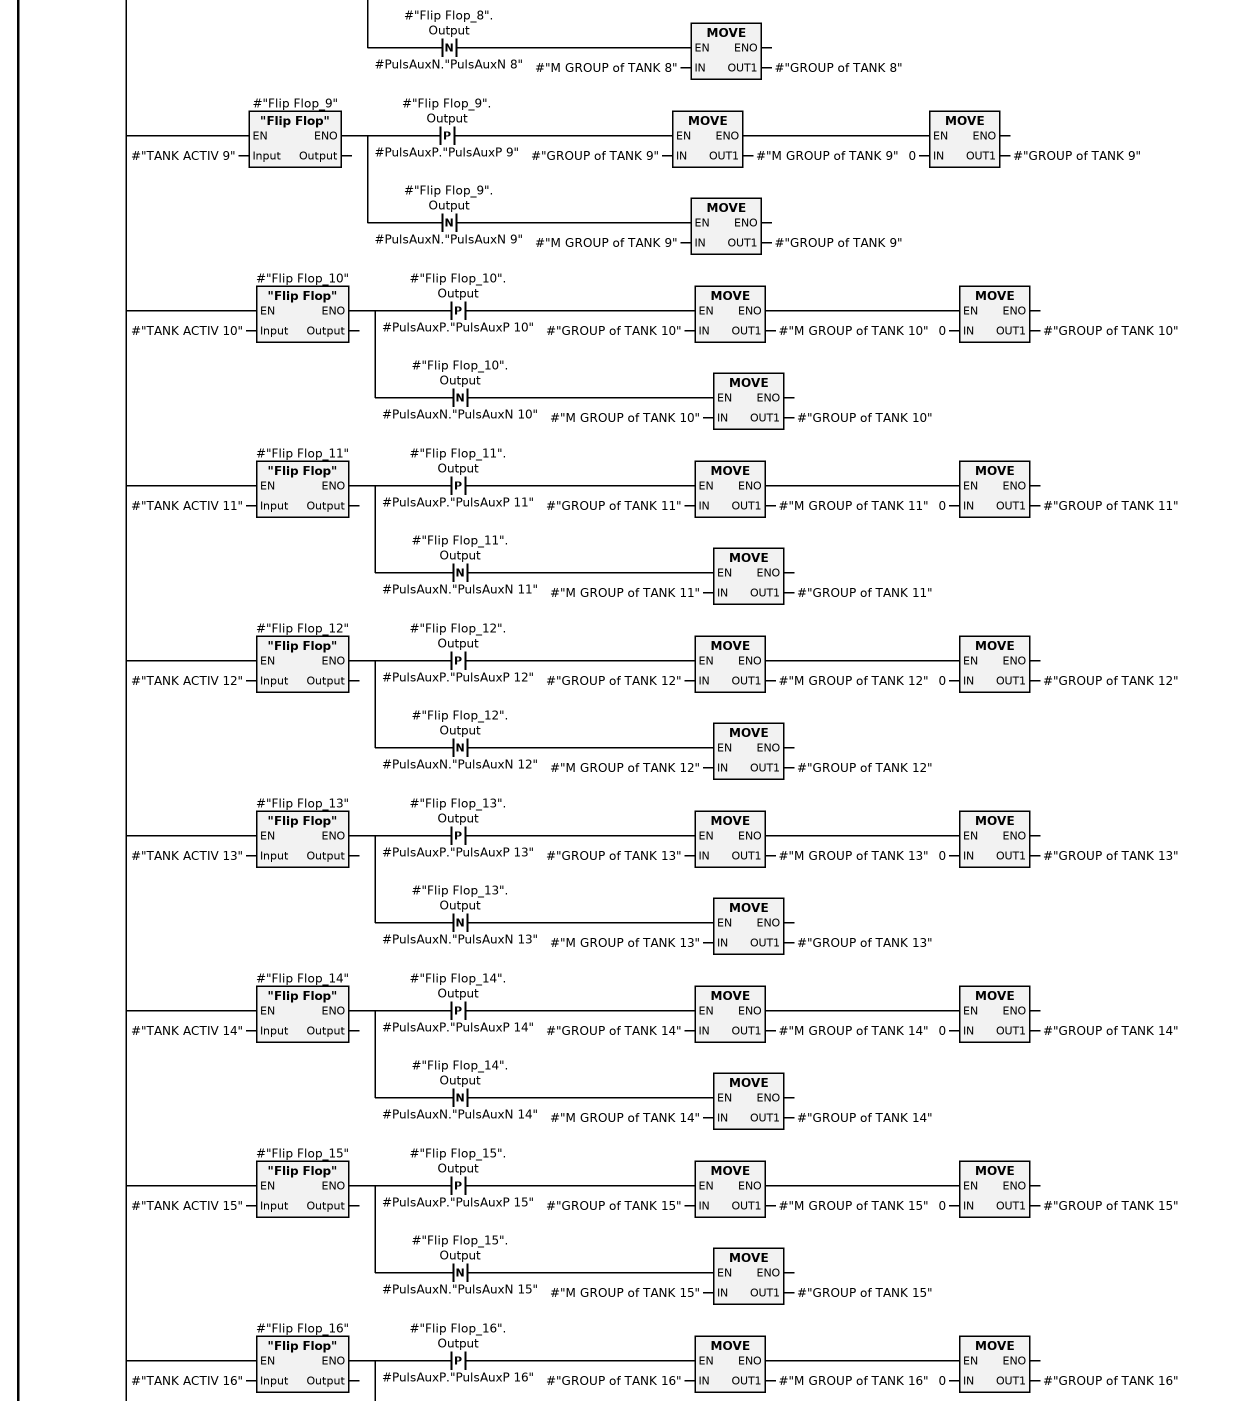
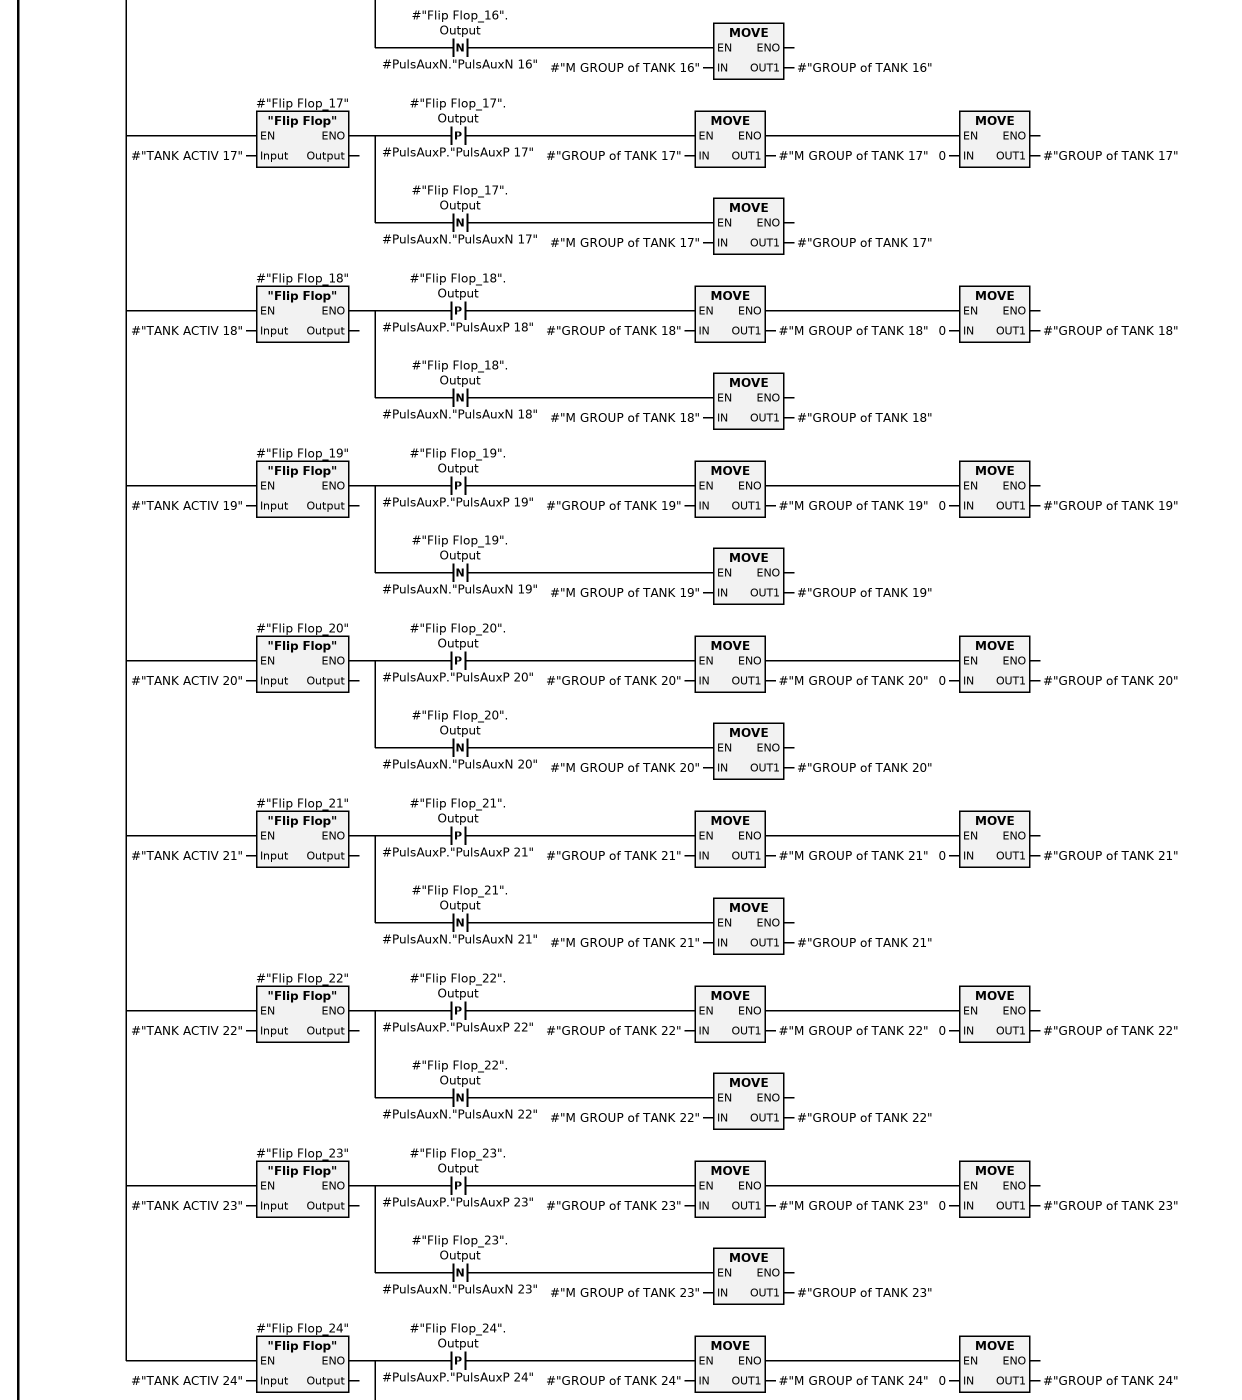
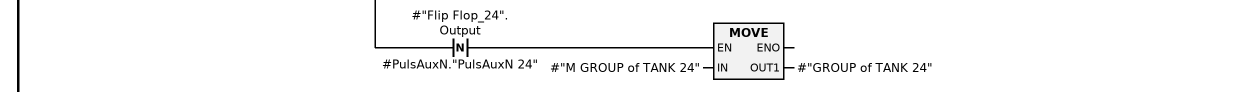
   RUNG wire#powerrail
      I_Contact( #SetGroupSR )
      wire#w1
      #"Flip Flop_1"(Input := #"TANK ACTIV 1", Output =>)
      wire#w2
      P_Contact(operand := #"Flip Flop_1".Output, bit := #PulsAuxP."PulsAuxP 1")
      Move(in := #"GROUP of TANK 1", out1 => #"M GROUP of TANK 1")
      Move(in := 0, out1 => #"GROUP of TANK 1")
   END_RUNG
   RUNG wire#w2
      N_Contact(operand := #"Flip Flop_1".Output, bit := #PulsAuxN."PulsAuxN 1")
      Move(in := #"M GROUP of TANK 1", out1 => #"GROUP of TANK 1")
   END_RUNG
   RUNG wire#w1
      #"Flip Flop_2"(Input := #"TANK ACTIV 2", Output =>)
      wire#w3
      P_Contact(operand := #"Flip Flop_2".Output, bit := #PulsAuxP."PulsAuxP 2")
      Move(in := #"GROUP of TANK 2", out1 => #"M GROUP of TANK 2")
      Move(in := 0, out1 => #"GROUP of TANK 2")
   END_RUNG
   RUNG wire#w3
      N_Contact(operand := #"Flip Flop_2".Output, bit := #PulsAuxN."PulsAuxN 2")
      Move(in := #"M GROUP of TANK 2", out1 => #"GROUP of TANK 2")
   END_RUNG
   RUNG wire#w1
      #"Flip Flop_3"(Input := #"TANK ACTIV 3", Output =>)
      wire#w4
      P_Contact(operand := #"Flip Flop_3".Output, bit := #PulsAuxP."PulsAuxP 3")
      Move(in := #"GROUP of TANK 3", out1 => #"M GROUP of TANK 3")
      Move(in := 0, out1 => #"GROUP of TANK 3")
   END_RUNG
   RUNG wire#w4
      N_Contact(operand := #"Flip Flop_3".Output, bit := #PulsAuxN."PulsAuxN 3")
      Move(in := #"M GROUP of TANK 3", out1 => #"GROUP of TANK 3")
   END_RUNG
   RUNG wire#w1
      #"Flip Flop_4"(Input := #"TANK ACTIV 4", Output =>)
      wire#w5
      P_Contact(operand := #"Flip Flop_4".Output, bit := #PulsAuxP."PulsAuxP 4")
      Move(in := #"GROUP of TANK 4", out1 => #"M GROUP of TANK 4")
      Move(in := 0, out1 => #"GROUP of TANK 4")
   END_RUNG
   RUNG wire#w5
      N_Contact(operand := #"Flip Flop_4".Output, bit := #PulsAuxN."PulsAuxN 4")
      Move(in := #"M GROUP of TANK 4", out1 => #"GROUP of TANK 4")
   END_RUNG
   RUNG wire#w1
      #"Flip Flop_5"(Input := #"TANK ACTIV 5", Output =>)
      wire#w6
      P_Contact(operand := #"Flip Flop_5".Output, bit := #PulsAuxP."PulsAuxP 5")
      Move(in := #"GROUP of TANK 5", out1 => #"M GROUP of TANK 5")
      Move(in := 0, out1 => #"GROUP of TANK 5")
   END_RUNG
   RUNG wire#w6
      N_Contact(operand := #"Flip Flop_5".Output, bit := #PulsAuxN."PulsAuxN 5")
      Move(in := #"M GROUP of TANK 5", out1 => #"GROUP of TANK 5")
   END_RUNG
   RUNG wire#w1
      #"Flip Flop_6"(Input := #"TANK ACTIV 6", Output =>)
      wire#w7
      P_Contact(operand := #"Flip Flop_6".Output, bit := #PulsAuxP."PulsAuxP 6")
      Move(in := #"GROUP of TANK 6", out1 => #"M GROUP of TANK 6")
      Move(in := 0, out1 => #"GROUP of TANK 6")
   END_RUNG
   RUNG wire#w7
      N_Contact(operand := #"Flip Flop_6".Output, bit := #PulsAuxN."PulsAuxN 6")
      Move(in := #"M GROUP of TANK 6", out1 => #"GROUP of TANK 6")
   END_RUNG
   RUNG wire#w1
      #"Flip Flop_7"(Input := #"TANK ACTIV 7", Output =>)
      wire#w8
      P_Contact(operand := #"Flip Flop_7".Output, bit := #PulsAuxP."PulsAuxP 7")
      Move(in := #"GROUP of TANK 7", out1 => #"M GROUP of TANK 7")
      Move(in := 0, out1 => #"GROUP of TANK 7")
   END_RUNG
   RUNG wire#w8
      N_Contact(operand := #"Flip Flop_7".Output, bit := #PulsAuxN."PulsAuxN 7")
      Move(in := #"M GROUP of TANK 7", out1 => #"GROUP of TANK 7")
   END_RUNG
   RUNG wire#w1
      #"Flip Flop_8"(Input := #"TANK ACTIV 8", Output =>)
      wire#w9
      P_Contact(operand := #"Flip Flop_8".Output, bit := #PulsAuxP."PulsAuxP 8")
      Move(in := #"GROUP of TANK 8", out1 => #"M GROUP of TANK 8")
      Move(in := 0, out1 => #"GROUP of TANK 8")
   END_RUNG
   RUNG wire#w9
      N_Contact(operand := #"Flip Flop_8".Output, bit := #PulsAuxN."PulsAuxN 8")
      Move(in := #"M GROUP of TANK 8", out1 => #"GROUP of TANK 8")
   END_RUNG
   RUNG wire#w1
      #"Flip Flop_9"(Input := #"TANK ACTIV 9", Output =>)
      wire#w10
      P_Contact(operand := #"Flip Flop_9".Output, bit := #PulsAuxP."PulsAuxP 9")
      Move(in := #"GROUP of TANK 9", out1 => #"M GROUP of TANK 9")
      Move(in := 0, out1 => #"GROUP of TANK 9")
   END_RUNG
   RUNG wire#w10
      N_Contact(operand := #"Flip Flop_9".Output, bit := #PulsAuxN."PulsAuxN 9")
      Move(in := #"M GROUP of TANK 9", out1 => #"GROUP of TANK 9")
   END_RUNG
   RUNG wire#w1
      #"Flip Flop_10"(Input := #"TANK ACTIV 10", Output =>)
      wire#w11
      P_Contact(operand := #"Flip Flop_10".Output, bit := #PulsAuxP."PulsAuxP 10")
      Move(in := #"GROUP of TANK 10", out1 => #"M GROUP of TANK 10")
      Move(in := 0, out1 => #"GROUP of TANK 10")
   END_RUNG
   RUNG wire#w11
      N_Contact(operand := #"Flip Flop_10".Output, bit := #PulsAuxN."PulsAuxN 10")
      Move(in := #"M GROUP of TANK 10", out1 => #"GROUP of TANK 10")
   END_RUNG
   RUNG wire#w1
      #"Flip Flop_11"(Input := #"TANK ACTIV 11", Output =>)
      wire#w12
      P_Contact(operand := #"Flip Flop_11".Output, bit := #PulsAuxP."PulsAuxP 11")
      Move(in := #"GROUP of TANK 11", out1 => #"M GROUP of TANK 11")
      Move(in := 0, out1 => #"GROUP of TANK 11")
   END_RUNG
   RUNG wire#w12
      N_Contact(operand := #"Flip Flop_11".Output, bit := #PulsAuxN."PulsAuxN 11")
      Move(in := #"M GROUP of TANK 11", out1 => #"GROUP of TANK 11")
   END_RUNG
   RUNG wire#w1
      #"Flip Flop_12"(Input := #"TANK ACTIV 12", Output =>)
      wire#w13
      P_Contact(operand := #"Flip Flop_12".Output, bit := #PulsAuxP."PulsAuxP 12")
      Move(in := #"GROUP of TANK 12", out1 => #"M GROUP of TANK 12")
      Move(in := 0, out1 => #"GROUP of TANK 12")
   END_RUNG
   RUNG wire#w13
      N_Contact(operand := #"Flip Flop_12".Output, bit := #PulsAuxN."PulsAuxN 12")
      Move(in := #"M GROUP of TANK 12", out1 => #"GROUP of TANK 12")
   END_RUNG
   RUNG wire#w1
      #"Flip Flop_13"(Input := #"TANK ACTIV 13", Output =>)
      wire#w14
      P_Contact(operand := #"Flip Flop_13".Output, bit := #PulsAuxP."PulsAuxP 13")
      Move(in := #"GROUP of TANK 13", out1 => #"M GROUP of TANK 13")
      Move(in := 0, out1 => #"GROUP of TANK 13")
   END_RUNG
   RUNG wire#w14
      N_Contact(operand := #"Flip Flop_13".Output, bit := #PulsAuxN."PulsAuxN 13")
      Move(in := #"M GROUP of TANK 13", out1 => #"GROUP of TANK 13")
   END_RUNG
   RUNG wire#w1
      #"Flip Flop_14"(Input := #"TANK ACTIV 14", Output =>)
      wire#w15
      P_Contact(operand := #"Flip Flop_14".Output, bit := #PulsAuxP."PulsAuxP 14")
      Move(in := #"GROUP of TANK 14", out1 => #"M GROUP of TANK 14")
      Move(in := 0, out1 => #"GROUP of TANK 14")
   END_RUNG
   RUNG wire#w15
      N_Contact(operand := #"Flip Flop_14".Output, bit := #PulsAuxN."PulsAuxN 14")
      Move(in := #"M GROUP of TANK 14", out1 => #"GROUP of TANK 14")
   END_RUNG
   RUNG wire#w1
      #"Flip Flop_15"(Input := #"TANK ACTIV 15", Output =>)
      wire#w16
      P_Contact(operand := #"Flip Flop_15".Output, bit := #PulsAuxP."PulsAuxP 15")
      Move(in := #"GROUP of TANK 15", out1 => #"M GROUP of TANK 15")
      Move(in := 0, out1 => #"GROUP of TANK 15")
   END_RUNG
   RUNG wire#w16
      N_Contact(operand := #"Flip Flop_15".Output, bit := #PulsAuxN."PulsAuxN 15")
      Move(in := #"M GROUP of TANK 15", out1 => #"GROUP of TANK 15")
   END_RUNG
   RUNG wire#w1
      #"Flip Flop_16"(Input := #"TANK ACTIV 16", Output =>)
      wire#w17
      P_Contact(operand := #"Flip Flop_16".Output, bit := #PulsAuxP."PulsAuxP 16")
      Move(in := #"GROUP of TANK 16", out1 => #"M GROUP of TANK 16")
      Move(in := 0, out1 => #"GROUP of TANK 16")
   END_RUNG
   RUNG wire#w17
      N_Contact(operand := #"Flip Flop_16".Output, bit := #PulsAuxN."PulsAuxN 16")
      Move(in := #"M GROUP of TANK 16", out1 => #"GROUP of TANK 16")
   END_RUNG
   RUNG wire#w1
      #"Flip Flop_17"(Input := #"TANK ACTIV 17", Output =>)
      wire#w18
      P_Contact(operand := #"Flip Flop_17".Output, bit := #PulsAuxP."PulsAuxP 17")
      Move(in := #"GROUP of TANK 17", out1 => #"M GROUP of TANK 17")
      Move(in := 0, out1 => #"GROUP of TANK 17")
   END_RUNG
   RUNG wire#w18
      N_Contact(operand := #"Flip Flop_17".Output, bit := #PulsAuxN."PulsAuxN 17")
      Move(in := #"M GROUP of TANK 17", out1 => #"GROUP of TANK 17")
   END_RUNG
   RUNG wire#w1
      #"Flip Flop_18"(Input := #"TANK ACTIV 18", Output =>)
      wire#w19
      P_Contact(operand := #"Flip Flop_18".Output, bit := #PulsAuxP."PulsAuxP 18")
      Move(in := #"GROUP of TANK 18", out1 => #"M GROUP of TANK 18")
      Move(in := 0, out1 => #"GROUP of TANK 18")
   END_RUNG
   RUNG wire#w19
      N_Contact(operand := #"Flip Flop_18".Output, bit := #PulsAuxN."PulsAuxN 18")
      Move(in := #"M GROUP of TANK 18", out1 => #"GROUP of TANK 18")
   END_RUNG
   RUNG wire#w1
      #"Flip Flop_19"(Input := #"TANK ACTIV 19", Output =>)
      wire#w20
      P_Contact(operand := #"Flip Flop_19".Output, bit := #PulsAuxP."PulsAuxP 19")
      Move(in := #"GROUP of TANK 19", out1 => #"M GROUP of TANK 19")
      Move(in := 0, out1 => #"GROUP of TANK 19")
   END_RUNG
   RUNG wire#w20
      N_Contact(operand := #"Flip Flop_19".Output, bit := #PulsAuxN."PulsAuxN 19")
      Move(in := #"M GROUP of TANK 19", out1 => #"GROUP of TANK 19")
   END_RUNG
   RUNG wire#w1
      #"Flip Flop_20"(Input := #"TANK ACTIV 20", Output =>)
      wire#w21
      P_Contact(operand := #"Flip Flop_20".Output, bit := #PulsAuxP."PulsAuxP 20")
      Move(in := #"GROUP of TANK 20", out1 => #"M GROUP of TANK 20")
      Move(in := 0, out1 => #"GROUP of TANK 20")
   END_RUNG
   RUNG wire#w21
      N_Contact(operand := #"Flip Flop_20".Output, bit := #PulsAuxN."PulsAuxN 20")
      Move(in := #"M GROUP of TANK 20", out1 => #"GROUP of TANK 20")
   END_RUNG
   RUNG wire#w1
      #"Flip Flop_21"(Input := #"TANK ACTIV 21", Output =>)
      wire#w22
      P_Contact(operand := #"Flip Flop_21".Output, bit := #PulsAuxP."PulsAuxP 21")
      Move(in := #"GROUP of TANK 21", out1 => #"M GROUP of TANK 21")
      Move(in := 0, out1 => #"GROUP of TANK 21")
   END_RUNG
   RUNG wire#w22
      N_Contact(operand := #"Flip Flop_21".Output, bit := #PulsAuxN."PulsAuxN 21")
      Move(in := #"M GROUP of TANK 21", out1 => #"GROUP of TANK 21")
   END_RUNG
   RUNG wire#w1
      #"Flip Flop_22"(Input := #"TANK ACTIV 22", Output =>)
      wire#w23
      P_Contact(operand := #"Flip Flop_22".Output, bit := #PulsAuxP."PulsAuxP 22")
      Move(in := #"GROUP of TANK 22", out1 => #"M GROUP of TANK 22")
      Move(in := 0, out1 => #"GROUP of TANK 22")
   END_RUNG
   RUNG wire#w23
      N_Contact(operand := #"Flip Flop_22".Output, bit := #PulsAuxN."PulsAuxN 22")
      Move(in := #"M GROUP of TANK 22", out1 => #"GROUP of TANK 22")
   END_RUNG
   RUNG wire#w1
      #"Flip Flop_23"(Input := #"TANK ACTIV 23", Output =>)
      wire#w24
      P_Contact(operand := #"Flip Flop_23".Output, bit := #PulsAuxP."PulsAuxP 23")
      Move(in := #"GROUP of TANK 23", out1 => #"M GROUP of TANK 23")
      Move(in := 0, out1 => #"GROUP of TANK 23")
   END_RUNG
   RUNG wire#w24
      N_Contact(operand := #"Flip Flop_23".Output, bit := #PulsAuxN."PulsAuxN 23")
      Move(in := #"M GROUP of TANK 23", out1 => #"GROUP of TANK 23")
   END_RUNG
   RUNG wire#w1
      #"Flip Flop_24"(Input := #"TANK ACTIV 24", Output =>)
      wire#w25
      P_Contact(operand := #"Flip Flop_24".Output, bit := #PulsAuxP."PulsAuxP 24")
      Move(in := #"GROUP of TANK 24", out1 => #"M GROUP of TANK 24")
      Move(in := 0, out1 => #"GROUP of TANK 24")
   END_RUNG
   RUNG wire#w25
      N_Contact(operand := #"Flip Flop_24".Output, bit := #PulsAuxN."PulsAuxN 24")
      Move(in := #"M GROUP of TANK 24", out1 => #"GROUP of TANK 24")
   END_RUNG
   // the same network as SCL:
   #"Flip Flop_1"(EN := NOT #SetGroupSR, Input := #"TANK ACTIV 1", ENO => #_w1);   // "Flip Flop"
   #_w2 := #_w1 AND #"Flip Flop_1".Output AND NOT #PulsAuxP."PulsAuxP 1";   // rising edge of #"Flip Flop_1".Output
   #PulsAuxP."PulsAuxP 1" := #"Flip Flop_1".Output;
   IF #_w2 THEN
       #"M GROUP of TANK 1" := #"GROUP of TANK 1";
       #"GROUP of TANK 1" := 0;
   END_IF;
   #_w3 := #_w1 AND NOT #"Flip Flop_1".Output AND #PulsAuxN."PulsAuxN 1";   // falling edge of #"Flip Flop_1".Output
   #PulsAuxN."PulsAuxN 1" := #"Flip Flop_1".Output;
   IF #_w3 THEN #"GROUP of TANK 1" := #"M GROUP of TANK 1"; END_IF;
   #"Flip Flop_2"(EN := NOT #SetGroupSR, Input := #"TANK ACTIV 2", ENO => #_w4);   // "Flip Flop"
   #_w5 := #_w4 AND #"Flip Flop_2".Output AND NOT #PulsAuxP."PulsAuxP 2";   // rising edge of #"Flip Flop_2".Output
   #PulsAuxP."PulsAuxP 2" := #"Flip Flop_2".Output;
   IF #_w5 THEN
       #"M GROUP of TANK 2" := #"GROUP of TANK 2";
       #"GROUP of TANK 2" := 0;
   END_IF;
   #_w6 := #_w4 AND NOT #"Flip Flop_2".Output AND #PulsAuxN."PulsAuxN 2";   // falling edge of #"Flip Flop_2".Output
   #PulsAuxN."PulsAuxN 2" := #"Flip Flop_2".Output;
   IF #_w6 THEN #"GROUP of TANK 2" := #"M GROUP of TANK 2"; END_IF;
   #"Flip Flop_3"(EN := NOT #SetGroupSR, Input := #"TANK ACTIV 3", ENO => #_w7);   // "Flip Flop"
   #_w8 := #_w7 AND #"Flip Flop_3".Output AND NOT #PulsAuxP."PulsAuxP 3";   // rising edge of #"Flip Flop_3".Output
   #PulsAuxP."PulsAuxP 3" := #"Flip Flop_3".Output;
   IF #_w8 THEN
       #"M GROUP of TANK 3" := #"GROUP of TANK 3";
       #"GROUP of TANK 3" := 0;
   END_IF;
   #_w9 := #_w7 AND NOT #"Flip Flop_3".Output AND #PulsAuxN."PulsAuxN 3";   // falling edge of #"Flip Flop_3".Output
   #PulsAuxN."PulsAuxN 3" := #"Flip Flop_3".Output;
   IF #_w9 THEN #"GROUP of TANK 3" := #"M GROUP of TANK 3"; END_IF;
   #"Flip Flop_4"(EN := NOT #SetGroupSR, Input := #"TANK ACTIV 4", ENO => #_w10);   // "Flip Flop"
   #_w11 := #_w10 AND #"Flip Flop_4".Output AND NOT #PulsAuxP."PulsAuxP 4";   // rising edge of #"Flip Flop_4".Output
   #PulsAuxP."PulsAuxP 4" := #"Flip Flop_4".Output;
   IF #_w11 THEN
       #"M GROUP of TANK 4" := #"GROUP of TANK 4";
       #"GROUP of TANK 4" := 0;
   END_IF;
   #_w12 := #_w10 AND NOT #"Flip Flop_4".Output AND #PulsAuxN."PulsAuxN 4";   // falling edge of #"Flip Flop_4".Output
   #PulsAuxN."PulsAuxN 4" := #"Flip Flop_4".Output;
   IF #_w12 THEN #"GROUP of TANK 4" := #"M GROUP of TANK 4"; END_IF;
   #"Flip Flop_5"(EN := NOT #SetGroupSR, Input := #"TANK ACTIV 5", ENO => #_w13);   // "Flip Flop"
   #_w14 := #_w13 AND #"Flip Flop_5".Output AND NOT #PulsAuxP."PulsAuxP 5";   // rising edge of #"Flip Flop_5".Output
   #PulsAuxP."PulsAuxP 5" := #"Flip Flop_5".Output;
   IF #_w14 THEN
       #"M GROUP of TANK 5" := #"GROUP of TANK 5";
       #"GROUP of TANK 5" := 0;
   END_IF;
   #_w15 := #_w13 AND NOT #"Flip Flop_5".Output AND #PulsAuxN."PulsAuxN 5";   // falling edge of #"Flip Flop_5".Output
   #PulsAuxN."PulsAuxN 5" := #"Flip Flop_5".Output;
   IF #_w15 THEN #"GROUP of TANK 5" := #"M GROUP of TANK 5"; END_IF;
   #"Flip Flop_6"(EN := NOT #SetGroupSR, Input := #"TANK ACTIV 6", ENO => #_w16);   // "Flip Flop"
   #_w17 := #_w16 AND #"Flip Flop_6".Output AND NOT #PulsAuxP."PulsAuxP 6";   // rising edge of #"Flip Flop_6".Output
   #PulsAuxP."PulsAuxP 6" := #"Flip Flop_6".Output;
   IF #_w17 THEN
       #"M GROUP of TANK 6" := #"GROUP of TANK 6";
       #"GROUP of TANK 6" := 0;
   END_IF;
   #_w18 := #_w16 AND NOT #"Flip Flop_6".Output AND #PulsAuxN."PulsAuxN 6";   // falling edge of #"Flip Flop_6".Output
   #PulsAuxN."PulsAuxN 6" := #"Flip Flop_6".Output;
   IF #_w18 THEN #"GROUP of TANK 6" := #"M GROUP of TANK 6"; END_IF;
   #"Flip Flop_7"(EN := NOT #SetGroupSR, Input := #"TANK ACTIV 7", ENO => #_w19);   // "Flip Flop"
   #_w20 := #_w19 AND #"Flip Flop_7".Output AND NOT #PulsAuxP."PulsAuxP 7";   // rising edge of #"Flip Flop_7".Output
   #PulsAuxP."PulsAuxP 7" := #"Flip Flop_7".Output;
   IF #_w20 THEN
       #"M GROUP of TANK 7" := #"GROUP of TANK 7";
       #"GROUP of TANK 7" := 0;
   END_IF;
   #_w21 := #_w19 AND NOT #"Flip Flop_7".Output AND #PulsAuxN."PulsAuxN 7";   // falling edge of #"Flip Flop_7".Output
   #PulsAuxN."PulsAuxN 7" := #"Flip Flop_7".Output;
   IF #_w21 THEN #"GROUP of TANK 7" := #"M GROUP of TANK 7"; END_IF;
   #"Flip Flop_8"(EN := NOT #SetGroupSR, Input := #"TANK ACTIV 8", ENO => #_w22);   // "Flip Flop"
   #_w23 := #_w22 AND #"Flip Flop_8".Output AND NOT #PulsAuxP."PulsAuxP 8";   // rising edge of #"Flip Flop_8".Output
   #PulsAuxP."PulsAuxP 8" := #"Flip Flop_8".Output;
   IF #_w23 THEN
       #"M GROUP of TANK 8" := #"GROUP of TANK 8";
       #"GROUP of TANK 8" := 0;
   END_IF;
   #_w24 := #_w22 AND NOT #"Flip Flop_8".Output AND #PulsAuxN."PulsAuxN 8";   // falling edge of #"Flip Flop_8".Output
   #PulsAuxN."PulsAuxN 8" := #"Flip Flop_8".Output;
   IF #_w24 THEN #"GROUP of TANK 8" := #"M GROUP of TANK 8"; END_IF;
   #"Flip Flop_9"(EN := NOT #SetGroupSR, Input := #"TANK ACTIV 9", ENO => #_w25);   // "Flip Flop"
   #_w26 := #_w25 AND #"Flip Flop_9".Output AND NOT #PulsAuxP."PulsAuxP 9";   // rising edge of #"Flip Flop_9".Output
   #PulsAuxP."PulsAuxP 9" := #"Flip Flop_9".Output;
   IF #_w26 THEN
       #"M GROUP of TANK 9" := #"GROUP of TANK 9";
       #"GROUP of TANK 9" := 0;
   END_IF;
   #_w27 := #_w25 AND NOT #"Flip Flop_9".Output AND #PulsAuxN."PulsAuxN 9";   // falling edge of #"Flip Flop_9".Output
   #PulsAuxN."PulsAuxN 9" := #"Flip Flop_9".Output;
   IF #_w27 THEN #"GROUP of TANK 9" := #"M GROUP of TANK 9"; END_IF;
   #"Flip Flop_10"(EN := NOT #SetGroupSR, Input := #"TANK ACTIV 10", ENO => #_w28);   // "Flip Flop"
   #_w29 := #_w28 AND #"Flip Flop_10".Output AND NOT #PulsAuxP."PulsAuxP 10";   // rising edge of #"Flip Flop_10".Output
   #PulsAuxP."PulsAuxP 10" := #"Flip Flop_10".Output;
   IF #_w29 THEN
       #"M GROUP of TANK 10" := #"GROUP of TANK 10";
       #"GROUP of TANK 10" := 0;
   END_IF;
   #_w30 := #_w28 AND NOT #"Flip Flop_10".Output AND #PulsAuxN."PulsAuxN 10";   // falling edge of #"Flip Flop_10".Output
   #PulsAuxN."PulsAuxN 10" := #"Flip Flop_10".Output;
   IF #_w30 THEN #"GROUP of TANK 10" := #"M GROUP of TANK 10"; END_IF;
   #"Flip Flop_11"(EN := NOT #SetGroupSR, Input := #"TANK ACTIV 11", ENO => #_w31);   // "Flip Flop"
   #_w32 := #_w31 AND #"Flip Flop_11".Output AND NOT #PulsAuxP."PulsAuxP 11";   // rising edge of #"Flip Flop_11".Output
   #PulsAuxP."PulsAuxP 11" := #"Flip Flop_11".Output;
   IF #_w32 THEN
       #"M GROUP of TANK 11" := #"GROUP of TANK 11";
       #"GROUP of TANK 11" := 0;
   END_IF;
   #_w33 := #_w31 AND NOT #"Flip Flop_11".Output AND #PulsAuxN."PulsAuxN 11";   // falling edge of #"Flip Flop_11".Output
   #PulsAuxN."PulsAuxN 11" := #"Flip Flop_11".Output;
   IF #_w33 THEN #"GROUP of TANK 11" := #"M GROUP of TANK 11"; END_IF;
   #"Flip Flop_12"(EN := NOT #SetGroupSR, Input := #"TANK ACTIV 12", ENO => #_w34);   // "Flip Flop"
   #_w35 := #_w34 AND #"Flip Flop_12".Output AND NOT #PulsAuxP."PulsAuxP 12";   // rising edge of #"Flip Flop_12".Output
   #PulsAuxP."PulsAuxP 12" := #"Flip Flop_12".Output;
   IF #_w35 THEN
       #"M GROUP of TANK 12" := #"GROUP of TANK 12";
       #"GROUP of TANK 12" := 0;
   END_IF;
   #_w36 := #_w34 AND NOT #"Flip Flop_12".Output AND #PulsAuxN."PulsAuxN 12";   // falling edge of #"Flip Flop_12".Output
   #PulsAuxN."PulsAuxN 12" := #"Flip Flop_12".Output;
   IF #_w36 THEN #"GROUP of TANK 12" := #"M GROUP of TANK 12"; END_IF;
   #"Flip Flop_13"(EN := NOT #SetGroupSR, Input := #"TANK ACTIV 13", ENO => #_w37);   // "Flip Flop"
   #_w38 := #_w37 AND #"Flip Flop_13".Output AND NOT #PulsAuxP."PulsAuxP 13";   // rising edge of #"Flip Flop_13".Output
   #PulsAuxP."PulsAuxP 13" := #"Flip Flop_13".Output;
   IF #_w38 THEN
       #"M GROUP of TANK 13" := #"GROUP of TANK 13";
       #"GROUP of TANK 13" := 0;
   END_IF;
   #_w39 := #_w37 AND NOT #"Flip Flop_13".Output AND #PulsAuxN."PulsAuxN 13";   // falling edge of #"Flip Flop_13".Output
   #PulsAuxN."PulsAuxN 13" := #"Flip Flop_13".Output;
   IF #_w39 THEN #"GROUP of TANK 13" := #"M GROUP of TANK 13"; END_IF;
   #"Flip Flop_14"(EN := NOT #SetGroupSR, Input := #"TANK ACTIV 14", ENO => #_w40);   // "Flip Flop"
   #_w41 := #_w40 AND #"Flip Flop_14".Output AND NOT #PulsAuxP."PulsAuxP 14";   // rising edge of #"Flip Flop_14".Output
   #PulsAuxP."PulsAuxP 14" := #"Flip Flop_14".Output;
   IF #_w41 THEN
       #"M GROUP of TANK 14" := #"GROUP of TANK 14";
       #"GROUP of TANK 14" := 0;
   END_IF;
   #_w42 := #_w40 AND NOT #"Flip Flop_14".Output AND #PulsAuxN."PulsAuxN 14";   // falling edge of #"Flip Flop_14".Output
   #PulsAuxN."PulsAuxN 14" := #"Flip Flop_14".Output;
   IF #_w42 THEN #"GROUP of TANK 14" := #"M GROUP of TANK 14"; END_IF;
   #"Flip Flop_15"(EN := NOT #SetGroupSR, Input := #"TANK ACTIV 15", ENO => #_w43);   // "Flip Flop"
   #_w44 := #_w43 AND #"Flip Flop_15".Output AND NOT #PulsAuxP."PulsAuxP 15";   // rising edge of #"Flip Flop_15".Output
   #PulsAuxP."PulsAuxP 15" := #"Flip Flop_15".Output;
   IF #_w44 THEN
       #"M GROUP of TANK 15" := #"GROUP of TANK 15";
       #"GROUP of TANK 15" := 0;
   END_IF;
   #_w45 := #_w43 AND NOT #"Flip Flop_15".Output AND #PulsAuxN."PulsAuxN 15";   // falling edge of #"Flip Flop_15".Output
   #PulsAuxN."PulsAuxN 15" := #"Flip Flop_15".Output;
   IF #_w45 THEN #"GROUP of TANK 15" := #"M GROUP of TANK 15"; END_IF;
   #"Flip Flop_16"(EN := NOT #SetGroupSR, Input := #"TANK ACTIV 16", ENO => #_w46);   // "Flip Flop"
   #_w47 := #_w46 AND #"Flip Flop_16".Output AND NOT #PulsAuxP."PulsAuxP 16";   // rising edge of #"Flip Flop_16".Output
   #PulsAuxP."PulsAuxP 16" := #"Flip Flop_16".Output;
   IF #_w47 THEN
       #"M GROUP of TANK 16" := #"GROUP of TANK 16";
       #"GROUP of TANK 16" := 0;
   END_IF;
   #_w48 := #_w46 AND NOT #"Flip Flop_16".Output AND #PulsAuxN."PulsAuxN 16";   // falling edge of #"Flip Flop_16".Output
   #PulsAuxN."PulsAuxN 16" := #"Flip Flop_16".Output;
   IF #_w48 THEN #"GROUP of TANK 16" := #"M GROUP of TANK 16"; END_IF;
   #"Flip Flop_17"(EN := NOT #SetGroupSR, Input := #"TANK ACTIV 17", ENO => #_w49);   // "Flip Flop"
   #_w50 := #_w49 AND #"Flip Flop_17".Output AND NOT #PulsAuxP."PulsAuxP 17";   // rising edge of #"Flip Flop_17".Output
   #PulsAuxP."PulsAuxP 17" := #"Flip Flop_17".Output;
   IF #_w50 THEN
       #"M GROUP of TANK 17" := #"GROUP of TANK 17";
       #"GROUP of TANK 17" := 0;
   END_IF;
   #_w51 := #_w49 AND NOT #"Flip Flop_17".Output AND #PulsAuxN."PulsAuxN 17";   // falling edge of #"Flip Flop_17".Output
   #PulsAuxN."PulsAuxN 17" := #"Flip Flop_17".Output;
   IF #_w51 THEN #"GROUP of TANK 17" := #"M GROUP of TANK 17"; END_IF;
   #"Flip Flop_18"(EN := NOT #SetGroupSR, Input := #"TANK ACTIV 18", ENO => #_w52);   // "Flip Flop"
   #_w53 := #_w52 AND #"Flip Flop_18".Output AND NOT #PulsAuxP."PulsAuxP 18";   // rising edge of #"Flip Flop_18".Output
   #PulsAuxP."PulsAuxP 18" := #"Flip Flop_18".Output;
   IF #_w53 THEN
       #"M GROUP of TANK 18" := #"GROUP of TANK 18";
       #"GROUP of TANK 18" := 0;
   END_IF;
   #_w54 := #_w52 AND NOT #"Flip Flop_18".Output AND #PulsAuxN."PulsAuxN 18";   // falling edge of #"Flip Flop_18".Output
   #PulsAuxN."PulsAuxN 18" := #"Flip Flop_18".Output;
   IF #_w54 THEN #"GROUP of TANK 18" := #"M GROUP of TANK 18"; END_IF;
   #"Flip Flop_19"(EN := NOT #SetGroupSR, Input := #"TANK ACTIV 19", ENO => #_w55);   // "Flip Flop"
   #_w56 := #_w55 AND #"Flip Flop_19".Output AND NOT #PulsAuxP."PulsAuxP 19";   // rising edge of #"Flip Flop_19".Output
   #PulsAuxP."PulsAuxP 19" := #"Flip Flop_19".Output;
   IF #_w56 THEN
       #"M GROUP of TANK 19" := #"GROUP of TANK 19";
       #"GROUP of TANK 19" := 0;
   END_IF;
   #_w57 := #_w55 AND NOT #"Flip Flop_19".Output AND #PulsAuxN."PulsAuxN 19";   // falling edge of #"Flip Flop_19".Output
   #PulsAuxN."PulsAuxN 19" := #"Flip Flop_19".Output;
   IF #_w57 THEN #"GROUP of TANK 19" := #"M GROUP of TANK 19"; END_IF;
   #"Flip Flop_20"(EN := NOT #SetGroupSR, Input := #"TANK ACTIV 20", ENO => #_w58);   // "Flip Flop"
   #_w59 := #_w58 AND #"Flip Flop_20".Output AND NOT #PulsAuxP."PulsAuxP 20";   // rising edge of #"Flip Flop_20".Output
   #PulsAuxP."PulsAuxP 20" := #"Flip Flop_20".Output;
   IF #_w59 THEN
       #"M GROUP of TANK 20" := #"GROUP of TANK 20";
       #"GROUP of TANK 20" := 0;
   END_IF;
   #_w60 := #_w58 AND NOT #"Flip Flop_20".Output AND #PulsAuxN."PulsAuxN 20";   // falling edge of #"Flip Flop_20".Output
   #PulsAuxN."PulsAuxN 20" := #"Flip Flop_20".Output;
   IF #_w60 THEN #"GROUP of TANK 20" := #"M GROUP of TANK 20"; END_IF;
   #"Flip Flop_21"(EN := NOT #SetGroupSR, Input := #"TANK ACTIV 21", ENO => #_w61);   // "Flip Flop"
   #_w62 := #_w61 AND #"Flip Flop_21".Output AND NOT #PulsAuxP."PulsAuxP 21";   // rising edge of #"Flip Flop_21".Output
   #PulsAuxP."PulsAuxP 21" := #"Flip Flop_21".Output;
   IF #_w62 THEN
       #"M GROUP of TANK 21" := #"GROUP of TANK 21";
       #"GROUP of TANK 21" := 0;
   END_IF;
   #_w63 := #_w61 AND NOT #"Flip Flop_21".Output AND #PulsAuxN."PulsAuxN 21";   // falling edge of #"Flip Flop_21".Output
   #PulsAuxN."PulsAuxN 21" := #"Flip Flop_21".Output;
   IF #_w63 THEN #"GROUP of TANK 21" := #"M GROUP of TANK 21"; END_IF;
   #"Flip Flop_22"(EN := NOT #SetGroupSR, Input := #"TANK ACTIV 22", ENO => #_w64);   // "Flip Flop"
   #_w65 := #_w64 AND #"Flip Flop_22".Output AND NOT #PulsAuxP."PulsAuxP 22";   // rising edge of #"Flip Flop_22".Output
   #PulsAuxP."PulsAuxP 22" := #"Flip Flop_22".Output;
   IF #_w65 THEN
       #"M GROUP of TANK 22" := #"GROUP of TANK 22";
       #"GROUP of TANK 22" := 0;
   END_IF;
   #_w66 := #_w64 AND NOT #"Flip Flop_22".Output AND #PulsAuxN."PulsAuxN 22";   // falling edge of #"Flip Flop_22".Output
   #PulsAuxN."PulsAuxN 22" := #"Flip Flop_22".Output;
   IF #_w66 THEN #"GROUP of TANK 22" := #"M GROUP of TANK 22"; END_IF;
   #"Flip Flop_23"(EN := NOT #SetGroupSR, Input := #"TANK ACTIV 23", ENO => #_w67);   // "Flip Flop"
   #_w68 := #_w67 AND #"Flip Flop_23".Output AND NOT #PulsAuxP."PulsAuxP 23";   // rising edge of #"Flip Flop_23".Output
   #PulsAuxP."PulsAuxP 23" := #"Flip Flop_23".Output;
   IF #_w68 THEN
       #"M GROUP of TANK 23" := #"GROUP of TANK 23";
       #"GROUP of TANK 23" := 0;
   END_IF;
   #_w69 := #_w67 AND NOT #"Flip Flop_23".Output AND #PulsAuxN."PulsAuxN 23";   // falling edge of #"Flip Flop_23".Output
   #PulsAuxN."PulsAuxN 23" := #"Flip Flop_23".Output;
   IF #_w69 THEN #"GROUP of TANK 23" := #"M GROUP of TANK 23"; END_IF;
   #"Flip Flop_24"(EN := NOT #SetGroupSR, Input := #"TANK ACTIV 24", ENO => #_w70);   // "Flip Flop"
   #_w71 := #_w70 AND #"Flip Flop_24".Output AND NOT #PulsAuxP."PulsAuxP 24";   // rising edge of #"Flip Flop_24".Output
   #PulsAuxP."PulsAuxP 24" := #"Flip Flop_24".Output;
   IF #_w71 THEN
       #"M GROUP of TANK 24" := #"GROUP of TANK 24";
       #"GROUP of TANK 24" := 0;
   END_IF;
   #_w72 := #_w70 AND NOT #"Flip Flop_24".Output AND #PulsAuxN."PulsAuxN 24";   // falling edge of #"Flip Flop_24".Output
   #PulsAuxN."PulsAuxN 24" := #"Flip Flop_24".Output;
   IF #_w72 THEN #"GROUP of TANK 24" := #"M GROUP of TANK 24"; END_IF;
END_REGION

REGION Network 36: GROUP ACTIVE SET
   // GROUP ACTIV to be used on HMI as SetTag on CLICK option